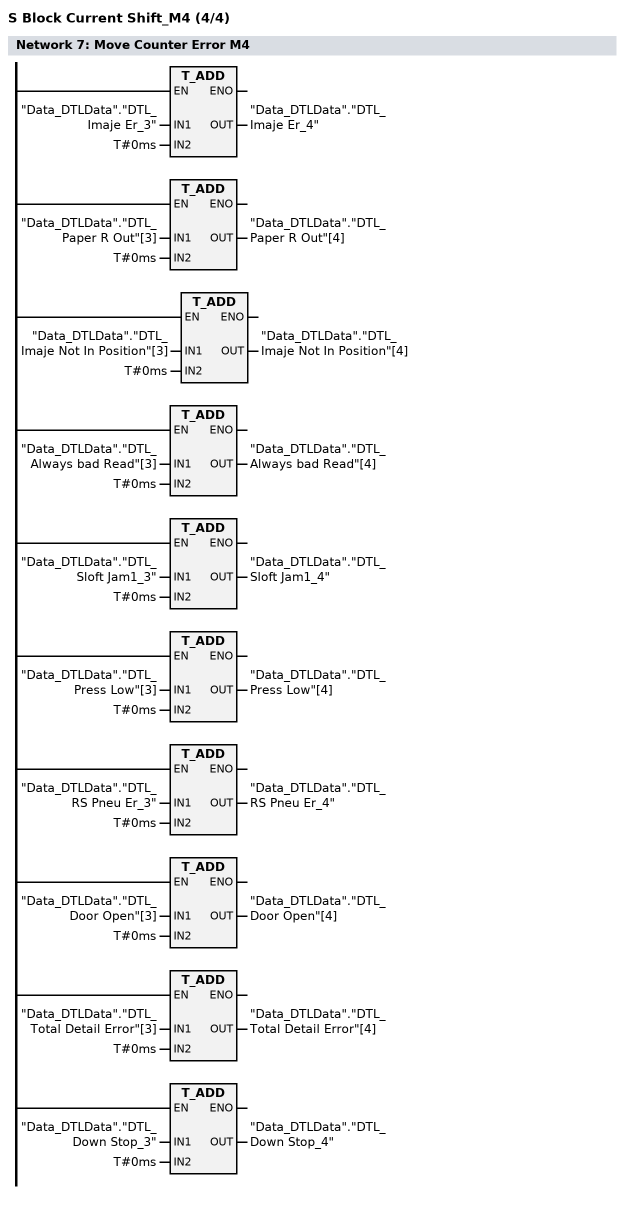
   "Data_DTLData"."DTL_Imaje Er_4" := T_ADD(IN1 := "Data_DTLData"."DTL_Imaje Er_3", IN2 := T#0ms);
   "Data_DTLData"."DTL_Paper R Out"[4] := T_ADD(IN1 := "Data_DTLData"."DTL_Paper R Out"[3], IN2 := T#0ms);
   "Data_DTLData"."DTL_Imaje Not In Position"[4] := T_ADD(IN1 := "Data_DTLData"."DTL_Imaje Not In Position"[3],
                           IN2 := T#0ms);
   "Data_DTLData"."DTL_Always bad Read"[4] := T_ADD(IN1 := "Data_DTLData"."DTL_Always bad Read"[3],
                           IN2 := T#0ms);
   "Data_DTLData"."DTL_Sloft Jam1_4" := T_ADD(IN1 := "Data_DTLData"."DTL_Sloft Jam1_3", IN2 := T#0ms);
   "Data_DTLData"."DTL_Press Low"[4] := T_ADD(IN1 := "Data_DTLData"."DTL_Press Low"[3], IN2 := T#0ms);
   "Data_DTLData"."DTL_RS Pneu Er_4" := T_ADD(IN1 := "Data_DTLData"."DTL_RS Pneu Er_3", IN2 := T#0ms);
   "Data_DTLData"."DTL_Door Open"[4] := T_ADD(IN1 := "Data_DTLData"."DTL_Door Open"[3], IN2 := T#0ms);
   "Data_DTLData"."DTL_Total Detail Error"[4] := T_ADD(IN1 := "Data_DTLData"."DTL_Total Detail Error"[3],
                           IN2 := T#0ms);
   "Data_DTLData"."DTL_Down Stop_4" := T_ADD(IN1 := "Data_DTLData"."DTL_Down Stop_3", IN2 := T#0ms);
END_REGION
END_FUNCTION_BLOCK

FUNCTION_BLOCK "S Block Current Shift_M5"   // FB14, LAD
{ S7_Optimized_Access := 'TRUE' }
VERSION : 0.1
BEGIN

REGION Network 1: Move Date Time M5
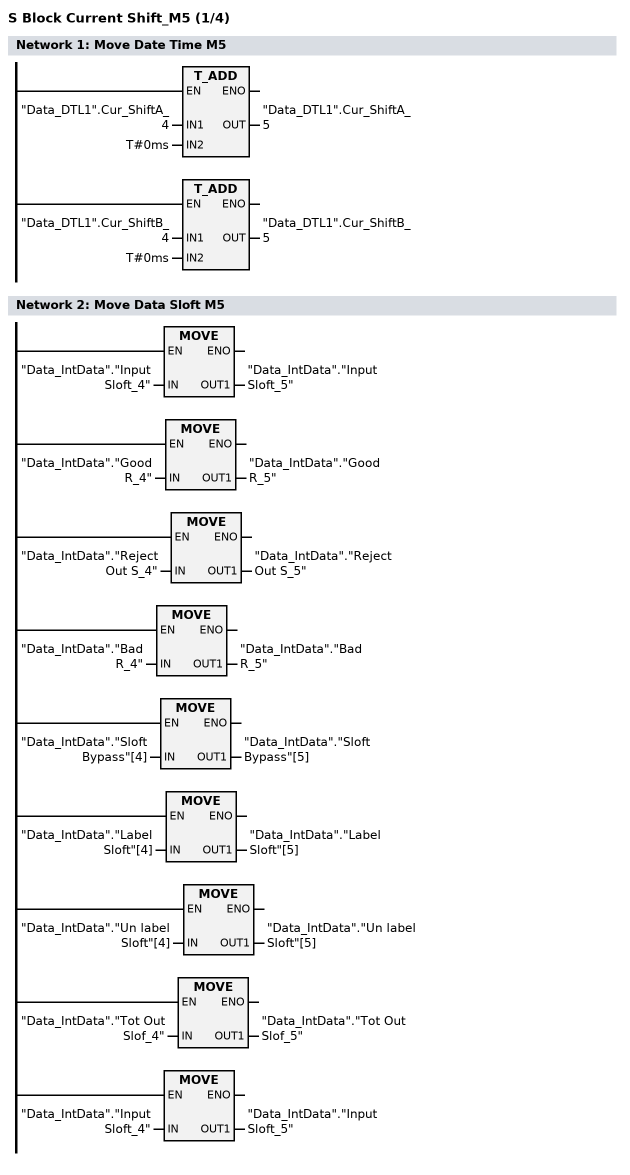
   "Data_DTL1".Cur_ShiftA_5 := T_ADD(IN1 := "Data_DTL1".Cur_ShiftA_4, IN2 := T#0ms);
   "Data_DTL1".Cur_ShiftB_5 := T_ADD(IN1 := "Data_DTL1".Cur_ShiftB_4, IN2 := T#0ms);
END_REGION

REGION Network 2: Move Data Sloft M5
   RUNG wire#powerrail
      { S7_GenerateENO := "TRUE" } Move(in := "Data_IntData"."Input Sloft_4", out1 => "Data_IntData"."Input Sloft_5")
   END_RUNG
   RUNG wire#powerrail
      { S7_GenerateENO := "TRUE" } Move(in := "Data_IntData"."Good R_4", out1 => "Data_IntData"."Good R_5")
   END_RUNG
   RUNG wire#powerrail
      { S7_GenerateENO := "TRUE" } Move(in := "Data_IntData"."Reject Out S_4", out1 => "Data_IntData"."Reject Out S_5")
   END_RUNG
   RUNG wire#powerrail
      { S7_GenerateENO := "TRUE" } Move(in := "Data_IntData"."Bad R_4", out1 => "Data_IntData"."Bad R_5")
   END_RUNG
   RUNG wire#powerrail
      { S7_GenerateENO := "TRUE" } Move(in := "Data_IntData"."Sloft Bypass"[4], out1 => "Data_IntData"."Sloft Bypass"[5])
   END_RUNG
   RUNG wire#powerrail
      { S7_GenerateENO := "TRUE" } Move(in := "Data_IntData"."Label Sloft"[4], out1 => "Data_IntData"."Label Sloft"[5])
   END_RUNG
   RUNG wire#powerrail
      { S7_GenerateENO := "TRUE" } Move(in := "Data_IntData"."Un label Sloft"[4], out1 => "Data_IntData"."Un label Sloft"[5])
   END_RUNG
   RUNG wire#powerrail
      { S7_GenerateENO := "TRUE" } Move(in := "Data_IntData"."Tot Out Slof_4", out1 => "Data_IntData"."Tot Out Slof_5")
   END_RUNG
   RUNG wire#powerrail
      { S7_GenerateENO := "TRUE" } Move(in := "Data_IntData"."Input Sloft_4", out1 => "Data_IntData"."Input Sloft_5")
   END_RUNG
   // the same network as SCL:
   "Data_IntData"."Input Sloft_5" := "Data_IntData"."Input Sloft_4";
   "Data_IntData"."Good R_5" := "Data_IntData"."Good R_4";
   "Data_IntData"."Reject Out S_5" := "Data_IntData"."Reject Out S_4";
   "Data_IntData"."Bad R_5" := "Data_IntData"."Bad R_4";
   "Data_IntData"."Sloft Bypass"[5] := "Data_IntData"."Sloft Bypass"[4];
   "Data_IntData"."Label Sloft"[5] := "Data_IntData"."Label Sloft"[4];
   "Data_IntData"."Un label Sloft"[5] := "Data_IntData"."Un label Sloft"[4];
   "Data_IntData"."Tot Out Slof_5" := "Data_IntData"."Tot Out Slof_4";
   "Data_IntData"."Input Sloft_5" := "Data_IntData"."Input Sloft_4";
END_REGION

REGION Network 3: Move Data Sloft Trigger & Aplicator M5
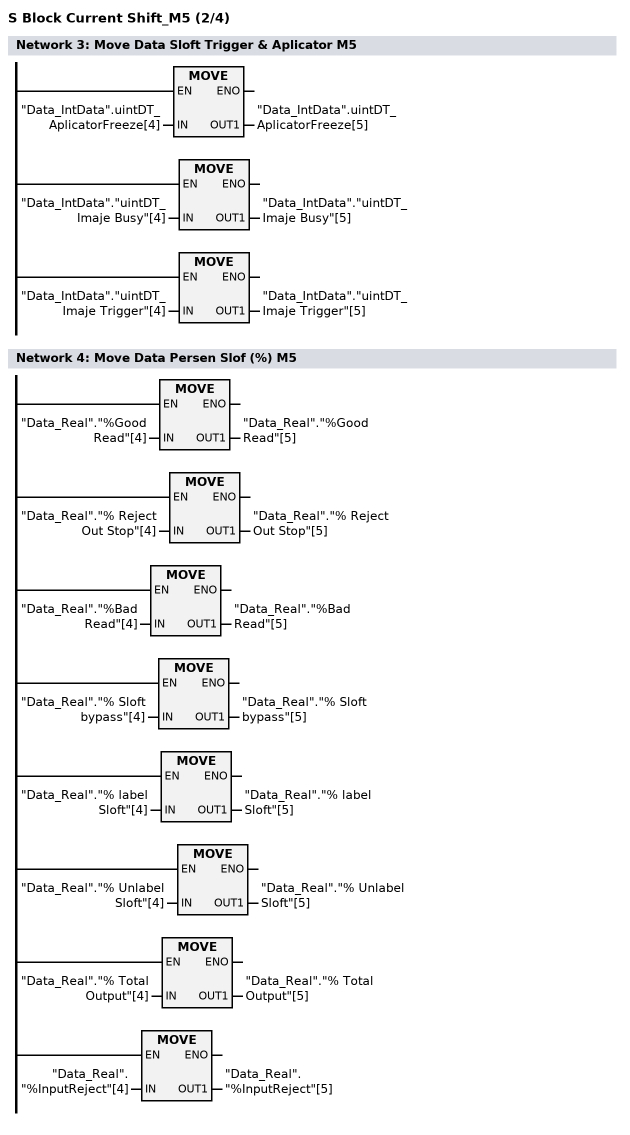
   RUNG wire#powerrail
      { S7_GenerateENO := "TRUE" } Move(in := "Data_IntData".uintDT_AplicatorFreeze[4], out1 => "Data_IntData".uintDT_AplicatorFreeze[5])
   END_RUNG
   RUNG wire#powerrail
      { S7_GenerateENO := "TRUE" } Move(in := "Data_IntData"."uintDT_Imaje Busy"[4], out1 => "Data_IntData"."uintDT_Imaje Busy"[5])
   END_RUNG
   RUNG wire#powerrail
      { S7_GenerateENO := "TRUE" } Move(in := "Data_IntData"."uintDT_Imaje Trigger"[4], out1 => "Data_IntData"."uintDT_Imaje Trigger"[5])
   END_RUNG
   // the same network as SCL:
   "Data_IntData".uintDT_AplicatorFreeze[5] := "Data_IntData".uintDT_AplicatorFreeze[4];
   "Data_IntData"."uintDT_Imaje Busy"[5] := "Data_IntData"."uintDT_Imaje Busy"[4];
   "Data_IntData"."uintDT_Imaje Trigger"[5] := "Data_IntData"."uintDT_Imaje Trigger"[4];
END_REGION

REGION Network 4: Move Data Persen Slof (%) M5
   RUNG wire#powerrail
      { S7_GenerateENO := "TRUE" } Move(in := "Data_Real"."%Good Read"[4], out1 => "Data_Real"."%Good Read"[5])
   END_RUNG
   RUNG wire#powerrail
      { S7_GenerateENO := "TRUE" } Move(in := "Data_Real"."% Reject Out Stop"[4], out1 => "Data_Real"."% Reject Out Stop"[5])
   END_RUNG
   RUNG wire#powerrail
      { S7_GenerateENO := "TRUE" } Move(in := "Data_Real"."%Bad Read"[4], out1 => "Data_Real"."%Bad Read"[5])
   END_RUNG
   RUNG wire#powerrail
      { S7_GenerateENO := "TRUE" } Move(in := "Data_Real"."% Sloft bypass"[4], out1 => "Data_Real"."% Sloft bypass"[5])
   END_RUNG
   RUNG wire#powerrail
      { S7_GenerateENO := "TRUE" } Move(in := "Data_Real"."% label Sloft"[4], out1 => "Data_Real"."% label Sloft"[5])
   END_RUNG
   RUNG wire#powerrail
      { S7_GenerateENO := "TRUE" } Move(in := "Data_Real"."% Unlabel Sloft"[4], out1 => "Data_Real"."% Unlabel Sloft"[5])
   END_RUNG
   RUNG wire#powerrail
      { S7_GenerateENO := "TRUE" } Move(in := "Data_Real"."% Total Output"[4], out1 => "Data_Real"."% Total Output"[5])
   END_RUNG
   RUNG wire#powerrail
      { S7_GenerateENO := "TRUE" } Move(in := "Data_Real"."%InputReject"[4], out1 => "Data_Real"."%InputReject"[5])
   END_RUNG
   // the same network as SCL:
   "Data_Real"."%Good Read"[5] := "Data_Real"."%Good Read"[4];
   "Data_Real"."% Reject Out Stop"[5] := "Data_Real"."% Reject Out Stop"[4];
   "Data_Real"."%Bad Read"[5] := "Data_Real"."%Bad Read"[4];
   "Data_Real"."% Sloft bypass"[5] := "Data_Real"."% Sloft bypass"[4];
   "Data_Real"."% label Sloft"[5] := "Data_Real"."% label Sloft"[4];
   "Data_Real"."% Unlabel Sloft"[5] := "Data_Real"."% Unlabel Sloft"[4];
   "Data_Real"."% Total Output"[5] := "Data_Real"."% Total Output"[4];
   "Data_Real"."%InputReject"[5] := "Data_Real"."%InputReject"[4];
END_REGION

REGION Network 5: Move Data Time Mesin M5
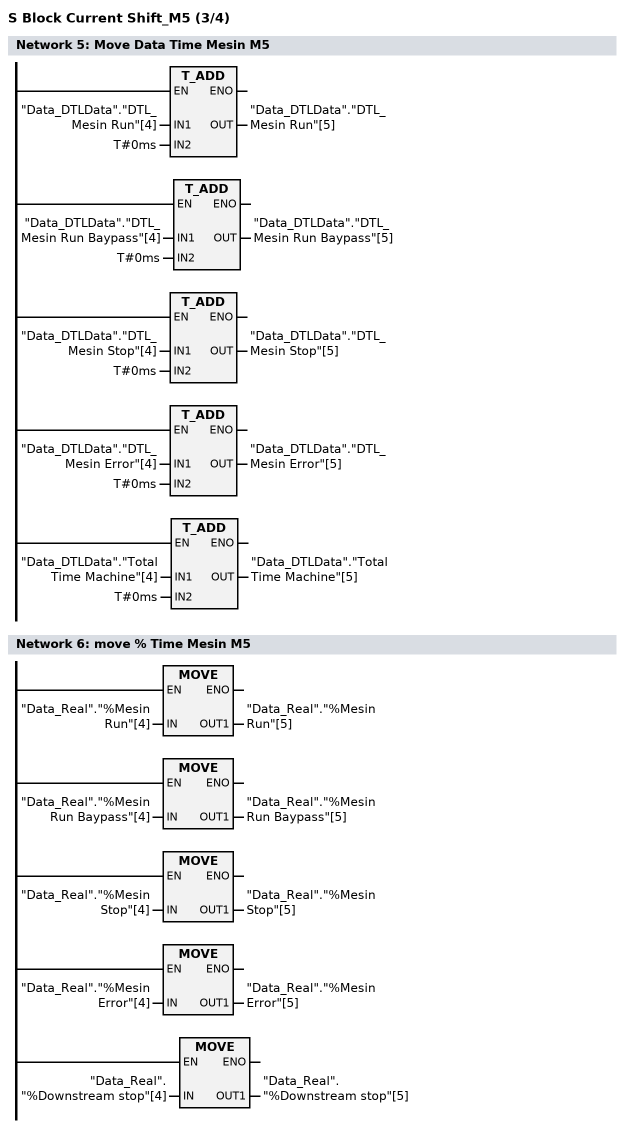
   "Data_DTLData"."DTL_Mesin Run"[5] := T_ADD(IN1 := "Data_DTLData"."DTL_Mesin Run"[4], IN2 := T#0ms);
   "Data_DTLData"."DTL_Mesin Run Baypass"[5] := T_ADD(IN1 := "Data_DTLData"."DTL_Mesin Run Baypass"[4],
                           IN2 := T#0ms);
   "Data_DTLData"."DTL_Mesin Stop"[5] := T_ADD(IN1 := "Data_DTLData"."DTL_Mesin Stop"[4], IN2 := T#0ms);
   "Data_DTLData"."DTL_Mesin Error"[5] := T_ADD(IN1 := "Data_DTLData"."DTL_Mesin Error"[4], IN2 := T#0ms);
   "Data_DTLData"."Total Time Machine"[5] := T_ADD(IN1 := "Data_DTLData"."Total Time Machine"[4], IN2 := T#0ms);
END_REGION

REGION Network 6: move % Time Mesin M5
   RUNG wire#powerrail
      { S7_GenerateENO := "TRUE" } Move(in := "Data_Real"."%Mesin Run"[4], out1 => "Data_Real"."%Mesin Run"[5])
   END_RUNG
   RUNG wire#powerrail
      { S7_GenerateENO := "TRUE" } Move(in := "Data_Real"."%Mesin Run Baypass"[4], out1 => "Data_Real"."%Mesin Run Baypass"[5])
   END_RUNG
   RUNG wire#powerrail
      { S7_GenerateENO := "TRUE" } Move(in := "Data_Real"."%Mesin Stop"[4], out1 => "Data_Real"."%Mesin Stop"[5])
   END_RUNG
   RUNG wire#powerrail
      { S7_GenerateENO := "TRUE" } Move(in := "Data_Real"."%Mesin Error"[4], out1 => "Data_Real"."%Mesin Error"[5])
   END_RUNG
   RUNG wire#powerrail
      { S7_GenerateENO := "TRUE" } Move(in := "Data_Real"."%Downstream stop"[4], out1 => "Data_Real"."%Downstream stop"[5])
   END_RUNG
   // the same network as SCL:
   "Data_Real"."%Mesin Run"[5] := "Data_Real"."%Mesin Run"[4];
   "Data_Real"."%Mesin Run Baypass"[5] := "Data_Real"."%Mesin Run Baypass"[4];
   "Data_Real"."%Mesin Stop"[5] := "Data_Real"."%Mesin Stop"[4];
   "Data_Real"."%Mesin Error"[5] := "Data_Real"."%Mesin Error"[4];
   "Data_Real"."%Downstream stop"[5] := "Data_Real"."%Downstream stop"[4];
END_REGION

REGION Network 7: Move Counter Error M5
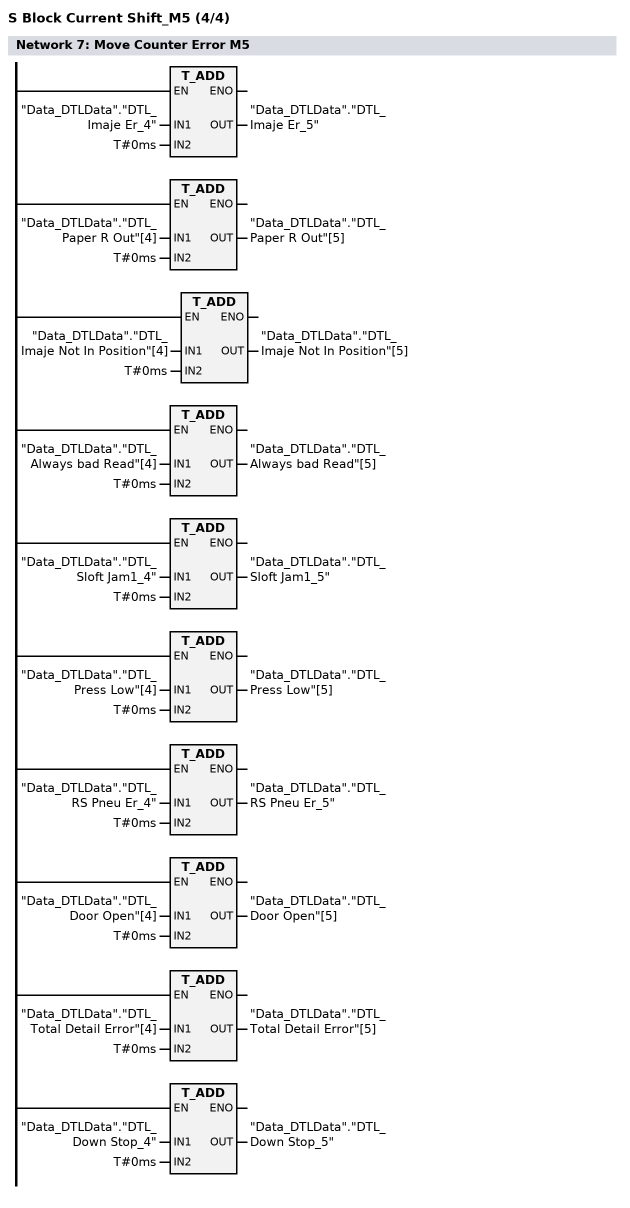
   "Data_DTLData"."DTL_Imaje Er_5" := T_ADD(IN1 := "Data_DTLData"."DTL_Imaje Er_4", IN2 := T#0ms);
   "Data_DTLData"."DTL_Paper R Out"[5] := T_ADD(IN1 := "Data_DTLData"."DTL_Paper R Out"[4], IN2 := T#0ms);
   "Data_DTLData"."DTL_Imaje Not In Position"[5] := T_ADD(IN1 := "Data_DTLData"."DTL_Imaje Not In Position"[4],
                           IN2 := T#0ms);
   "Data_DTLData"."DTL_Always bad Read"[5] := T_ADD(IN1 := "Data_DTLData"."DTL_Always bad Read"[4],
                           IN2 := T#0ms);
   "Data_DTLData"."DTL_Sloft Jam1_5" := T_ADD(IN1 := "Data_DTLData"."DTL_Sloft Jam1_4", IN2 := T#0ms);
   "Data_DTLData"."DTL_Press Low"[5] := T_ADD(IN1 := "Data_DTLData"."DTL_Press Low"[4], IN2 := T#0ms);
   "Data_DTLData"."DTL_RS Pneu Er_5" := T_ADD(IN1 := "Data_DTLData"."DTL_RS Pneu Er_4", IN2 := T#0ms);
   "Data_DTLData"."DTL_Door Open"[5] := T_ADD(IN1 := "Data_DTLData"."DTL_Door Open"[4], IN2 := T#0ms);
   "Data_DTLData"."DTL_Total Detail Error"[5] := T_ADD(IN1 := "Data_DTLData"."DTL_Total Detail Error"[4],
                           IN2 := T#0ms);
   "Data_DTLData"."DTL_Down Stop_5" := T_ADD(IN1 := "Data_DTLData"."DTL_Down Stop_4", IN2 := T#0ms);
END_REGION
END_FUNCTION_BLOCK

FUNCTION_BLOCK "AddReject2"   // FB15, SCL
{ S7_Optimized_Access := 'TRUE' }
VERSION : 0.1
   VAR_INPUT
      Sensor1 : Bool;
      Sensor2 : Bool;
      Sensor3 : Bool;
      Reedswicth1 : Bool;
      Reedswicth2 : Bool;
      BypassRS_AddRej : Bool;
      BypassRS_All_RS : Bool;
      PT_Timer_S1On : Time;
      PT_Timer_S1Off : Time;
      PT_Timer_S2On : Time;
      PT_Timer_S2Off : Time;
      PT_Timer_S3On : Time;
      PT_Timer_S3Off : Time;
      PT_Timer_DelayReject : Time;
      PT_Timer_DelayNonReject : Time;
   END_VAR
   VAR_OUTPUT
      Pneumatic1 : Bool;
      Pneumatic2 : Bool;
      Countaddrej : Time;
   END_VAR
   VAR
      SeqIndexReject : UInt;
      SeqIndexNonReject : UInt;
      FlagReject : Bool;
      FlagNonReject : Bool;
      FlagPneumatic : Bool;
      FlagSensor1 : Bool;
      FlagSensor2 : Bool;
      FlagSensor3 : Bool;
      FlagRS1Advance : Bool;
      FlagRS2Retract : Bool;
      RS1AdvanceError : Bool;
      RS2RetractError : Bool;
      AllRSAddRejectError : Bool;
      CountStop : Bool;
      InTimerDelayReject : Bool;
      InTimerDelaynonReject : Bool;
      InTimerErrorReject : Bool;
      InTimerErrorNonReject : Bool;
      InTimerRS1Error : Bool;
      InTimerRS2Error : Bool;
      R_TRIG_AddRejPSN1 : R_TRIG;
      F_TRIG_AddRejPSN1 : F_TRIG;
   END_VAR
BEGIN
   //Sensor 1
   "ttM_TimerAddRej1".TON(IN := #Sensor1,
                          PT := #PT_Timer_S1On);
   "tTM_TimerAddRej2".TON(IN := NOT #Sensor1,
                          PT := #PT_Timer_S1Off);
   IF "ttM_TimerAddRej1".Q THEN
       #FlagSensor1 := TRUE;
   END_IF;
   IF "tTM_TimerAddRej2".Q THEN
       #FlagSensor1 := FALSE;
   END_IF;

   //Sensor 2
   "tTM_TimerAddRej3".TON(IN := #Sensor2,
                          PT := #PT_Timer_S2On);
   "tTM_TimerAddRej4".TON(IN := NOT #Sensor2,
                          PT := #PT_Timer_S2Off);
   IF "tTM_TimerAddRej3".Q THEN
       #FlagSensor2 := TRUE;
   END_IF;
   IF "tTM_TimerAddRej4".Q THEN
       #FlagSensor2 := FALSE;
   END_IF;

   //Sensor 3
   "tTM_TimerAddRej5".TON(IN := #Sensor3,
                          PT := #PT_Timer_S3On);
   "tTM_TimerAddRej6".TON(IN := NOT #Sensor3,
                          PT := #PT_Timer_S3Off);
   IF "tTM_TimerAddRej5".Q THEN
       #FlagSensor3 := TRUE;
   END_IF;
   IF "tTM_TimerAddRej6".Q THEN
       #FlagSensor3 := FALSE;
   END_IF;

   //Reedswicth
   "tTM_TimerRS1_Adv".TON(IN := #InTimerRS1Error,
                          PT := T#1700ms);
   "tTM_TimerRS2_Ret".TON(IN := #InTimerRS2Error,
                          PT := T#1700ms);
   IF NOT #BypassRS_AddRej AND NOT #BypassRS_All_RS THEN
       //ReedSwicth Advance
       IF NOT #Pneumatic1 THEN
           #InTimerRS1Error := TRUE;
           "R_TRIG_RS1_Adv"(CLK := #Reedswicth1);
           IF #Reedswicth1 OR "R_TRIG_RS1_Adv".Q THEN
               #FlagRS1Advance := TRUE;
               #FlagRS2Retract := FALSE;
               #RS1AdvanceError := FALSE;
               #RS2RetractError := FALSE;
           ELSIF "tTM_TimerRS1_Adv".Q AND NOT #FlagRS1Advance THEN
               #FlagRS1Advance := FALSE;
               #FlagRS2Retract := FALSE;
               #RS1AdvanceError := TRUE;
               #RS2RetractError := FALSE;
           END_IF;
       ELSE
           #InTimerRS1Error := FALSE;
       END_IF;
       //ReeedSwicth Retract
       IF #Pneumatic2 THEN
           #InTimerRS2Error := TRUE;
           "R_TRIG_RS2_Ret"(CLK := #Reedswicth2);
           IF #Reedswicth2 OR "R_TRIG_RS2_Ret".Q THEN
               #FlagRS1Advance := FALSE;
               #FlagRS2Retract := TRUE;
               #RS1AdvanceError := FALSE;
               #RS2RetractError := FALSE;
           ELSIF "tTM_TimerRS2_Ret".Q AND NOT #FlagRS2Retract THEN
               #FlagRS1Advance := FALSE;
               #FlagRS2Retract := FALSE;
               #RS1AdvanceError := FALSE;
               #RS2RetractError := TRUE;
           END_IF;
       ELSE
           #InTimerRS2Error := FALSE;
       END_IF;
       //Error All ReedSwicth
       IF NOT #FlagRS1Advance AND NOT #FlagRS2Retract THEN
           "tTM_ErrorAllRSAddReject".TON(IN:=NOT #FlagRS1Advance AND NOT #FlagRS2Retract,
                                         PT:=T#3500ms);
           IF "tTM_ErrorAllRSAddReject".Q THEN
               IF #FlagSensor1 THEN
                   #Pneumatic1 := TRUE;
                   #Pneumatic2 := TRUE;
               ELSE
                   #Pneumatic1 := FALSE;
                   #Pneumatic2 := FALSE;
               END_IF;
               #AllRSAddRejectError := TRUE;
               #SeqIndexReject := 0;
               #SeqIndexNonReject := 0;
           END_IF;
       ELSE
           #AllRSAddRejectError := FALSE;
           "F_TRIG_AllRSAddrejError"(CLK:=#AllRSAddRejectError);
           IF "F_TRIG_AllRSAddrejError".Q THEN
               #SeqIndexReject := 1;
               #SeqIndexNonReject := 1;
           END_IF;
       END_IF;
   END_IF;

   //Reject Active
   IF #FlagSensor1 THEN
       IF NOT #AllRSAddRejectError THEN
           #SeqIndexNonReject := 1;
       END_IF;
       "tTM_DelayReject".TON(IN := #InTimerDelayReject,
                             PT := #PT_Timer_DelayReject);
       "tTM_ErrorReject".TON(IN := #InTimerErrorReject,
                             PT := T#2000ms);
       CASE #SeqIndexReject OF
           1:
               #InTimerErrorReject := FALSE;
               IF NOT #FlagSensor2 THEN
                   #Pneumatic1 := FALSE;
                   #Pneumatic2 := FALSE;
                   #SeqIndexReject := 10;
               ELSIF #FlagSensor2 THEN
                   IF "tTM_DelayReject".Q THEN
                       #Pneumatic1 := FALSE;
                       #Pneumatic2 := FALSE;
                       #SeqIndexReject := 10;
                   ELSE
                       #InTimerDelayReject := TRUE;
                   END_IF;
               END_IF;
           10:
               #InTimerDelayReject := FALSE;
               IF NOT #BypassRS_AddRej AND NOT #BypassRS_All_RS THEN
                   #SeqIndexReject := 20;
               ELSE
                   #SeqIndexReject := 1;
               END_IF;
           20:
               IF #FlagRS1Advance THEN
                   #SeqIndexReject := 1;
               ELSIF #RS1AdvanceError THEN
                   #Pneumatic1 := TRUE;
                   #Pneumatic2 := TRUE;
                   IF "tTM_ErrorReject".Q THEN
                       #SeqIndexReject := 1;
                   ELSE
                       #InTimerErrorReject := TRUE;
                   END_IF;
               END_IF;
           ELSE
               IF NOT #BypassRS_AddRej AND NOT #BypassRS_All_RS AND NOT #AllRSAddRejectError  THEN
                   #SeqIndexReject := 1;
               ELSE
                   #SeqIndexReject := 1;
               END_IF;
       END_CASE;
   END_IF;

   //Reject Start Non Active 
   IF NOT #FlagSensor1  THEN
       IF NOT #AllRSAddRejectError THEN
           #SeqIndexReject := 1;
       END_IF;
       "tTM_DelayNonReject".TON(IN := #InTimerDelaynonReject,
                                PT := #PT_Timer_DelayNonReject);
       "tTM_ErrorNonReject".TON(IN := #InTimerErrorNonReject,
                                PT := T#2000ms);
       CASE #SeqIndexNonReject OF
           1:
               #InTimerErrorNonReject := FALSE;
               IF NOT #FlagSensor3 THEN
                   #Pneumatic1 := TRUE;
                   #Pneumatic2 := TRUE;
                   #SeqIndexNonReject := 10;
               ELSIF #FlagSensor3 THEN
                   IF "tTM_DelayNonReject".Q THEN
                       #Pneumatic1 := TRUE;
                       #Pneumatic2 := TRUE;
                       #SeqIndexNonReject := 10;
                   ELSE
                       #InTimerDelaynonReject := TRUE;
                   END_IF;
               END_IF;
           10:
               #InTimerDelaynonReject := FALSE;
               IF NOT #BypassRS_AddRej AND NOT #BypassRS_All_RS THEN
                   #SeqIndexNonReject := 20;
               ELSE
                   #SeqIndexNonReject := 1;
               END_IF;
           20:
               IF #FlagRS2Retract THEN
                   #SeqIndexNonReject := 1;
               ELSIF #RS2RetractError THEN
                   #Pneumatic1 := FALSE;
                   #Pneumatic2 := FALSE;
                   IF "tTM_ErrorNonReject".Q THEN
                       #SeqIndexNonReject := 1;
                   ELSE
                       #InTimerErrorNonReject := TRUE;
                   END_IF;
               END_IF;
           ELSE
               IF NOT #BypassRS_AddRej AND NOT #BypassRS_All_RS AND NOT #AllRSAddRejectError THEN
                   #SeqIndexNonReject := 1;
               ELSE
                   #SeqIndexNonReject := 1;
               END_IF;
       END_CASE;
   END_IF;

   #R_TRIG_AddRejPSN1(CLK:=#FlagSensor1);
   #F_TRIG_AddRejPSN1(CLK:=#FlagSensor1);
   IF NOT #AllRSAddRejectError THEN
       IF #R_TRIG_AddRejPSN1.Q THEN
           #SeqIndexReject := 1;
       END_IF;
       IF #F_TRIG_AddRejPSN1.Q THEN
           #SeqIndexNonReject := 1;
       END_IF;
   END_IF;

   "tTM_CountAddReject".TON(IN:=#Sensor1,
                            PT:=T#5000ms);
   IF "tTM_CountAddReject".ET <>T#0ms THEN
       #Countaddrej :="tTM_CountAddReject".ET;
   ELSIF #CountStop THEN
       #Countaddrej := T#0ms;
   END_IF;


   //Error All ReedSwicth

   //Reject Active
   (*IF #FlagSensor1 THEN
     IF NOT #FlagSensor2 THEN
       #Pneumatic1 := FALSE;
       #Pneumatic2 := FALSE;
       #FlagPneumatic := FALSE;
     END_IF;
   END_IF;
   //Reject Start Non Active 
   IF NOT #FlagSensor1 THEN
       IF NOT #FlagSensor3 THEN
           #Pneumatic1 := TRUE;
           #Pneumatic2 := TRUE;
           #FlagPneumatic := TRUE;
       END_IF;
   END_IF;

   CASE #SeqIndex OF
       0:
           #RS1Error := FALSE;
           #RS2Error := FALSE;
           //Reject Start Active
           IF #FlagSensor1 AND NOT #RejectActive THEN
               #SeqIndex := 5;
           END_IF;
           //Reject Start Non Active 
           IF NOT #FlagSensor1 AND #RejectActive THEN
               #SeqIndex := 10;
           END_IF;
       5: //Reject Active
           IF NOT #FlagSensor2 THEN
               #Pneumatic1 := FALSE;
               #Pneumatic2 := FALSE;
               #FlagPneumatic := FALSE;
               #SeqIndex := 15;
           END_IF;
       10: //Reject Non Active
           IF NOT #FlagSensor3 THEN
               #Pneumatic1 := TRUE;
               #Pneumatic2 := TRUE;
               #FlagPneumatic := TRUE;
               #SeqIndex := 20;
           END_IF;
       15: // Active Finish
           IF #BypassRS_AddRej OR #BypassRS_All_RS THEN
               #RejectActive := TRUE;
               #SeqIndex := 0;
           ELSIF NOT #BypassRS_AddRej AND NOT #BypassRS_All_RS THEN
               IF #FlagRS1 THEN
                   #RejectActive := TRUE;
                   #SeqIndex := 0;
               ELSIF #RS1Error THEN
                   #Pneumatic1 := TRUE;
                   #Pneumatic2 := TRUE;
                   #FlagPneumatic := TRUE;
                   #RejectActive := FALSE;
                   #SeqIndex := 0;
               END_IF;
           END_IF;
       20: //Cek Non Active Finish
           IF #BypassRS_AddRej OR #BypassRS_All_RS THEN
               #RejectActive := FALSE;
               #SeqIndex := 0;
           ELSIF NOT #BypassRS_AddRej AND NOT #BypassRS_All_RS THEN
               IF #FlagRS2 THEN
                   #RejectActive := FALSE;
                   #SeqIndex := 0;
               ELSIF #RS2Error THEN
                   #Pneumatic1 := FALSE;
                   #Pneumatic2 := FALSE;
                   #FlagPneumatic := FALSE;
                   #RejectActive := TRUE;
                   #SeqIndex := 0;
               END_IF;
           END_IF;
       END_CASE;*)
END_FUNCTION_BLOCK

FUNCTION "RS 1 Pneumatic Pusher Advance" : Void   // FC1, LAD
{ S7_Optimized_Access := 'TRUE' }
VERSION : 0.1
BEGIN

REGION Network 1: Reed Switch Pneumatic 1 Advance Ready
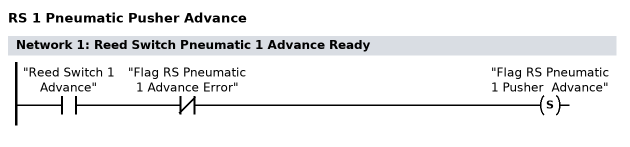
   RUNG wire#powerrail
      Contact( "Reed Switch 1 Advance" )
      I_Contact( "Flag RS Pneumatic 1 Advance Error" )
      S_Coil( "Flag RS Pneumatic 1 Pusher  Advance" )
   END_RUNG
   // the same network as SCL:
   IF "Reed Switch 1 Advance" AND NOT "Flag RS Pneumatic 1 Advance Error" THEN
       "Flag RS Pneumatic 1 Pusher  Advance" := TRUE;
   END_IF;
END_REGION
END_FUNCTION

FUNCTION "RS 2 Pneumatic Pusher Retract" : Void   // FC2, LAD
{ S7_Optimized_Access := 'TRUE' }
VERSION : 0.1
BEGIN

REGION Network 1: Reed Switch Pneumatic 1 Upper Ready
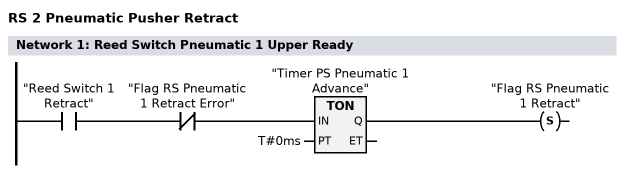
   "Timer PS Pneumatic 1 Advance".TON(IN := "Reed Switch 1 Retract" AND NOT "Flag RS Pneumatic 1 Retract Error",
                           PT := T#0ms);
   IF "Timer PS Pneumatic 1 Advance".Q THEN "Flag RS Pneumatic 1 Retract" := TRUE; END_IF;
END_REGION
END_FUNCTION

FUNCTION "RS 3 Pneumatic 3 Up" : Void   // FC3, LAD
{ S7_Optimized_Access := 'TRUE' }
VERSION : 0.1
BEGIN

REGION Network 1: Reed Switch Pneumatic 3 Up Ready
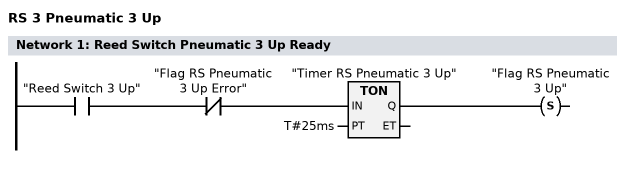
   "Timer RS Pneumatic 3 Up".TON(IN := "Reed Switch 3 Up" AND NOT "Flag RS Pneumatic 3 Up Error", PT := T#25ms);
   IF "Timer RS Pneumatic 3 Up".Q THEN "Flag RS Pneumatic 3 Up" := TRUE; END_IF;
END_REGION
END_FUNCTION

FUNCTION "RS 4 Pneumatic 3 Down" : Void   // FC4, LAD
{ S7_Optimized_Access := 'TRUE' }
VERSION : 0.1
BEGIN

REGION Network 1: Reed Switch Pneumatic 3 Down Ready
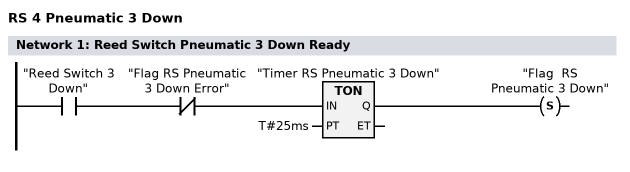
   "Timer RS Pneumatic 3 Down".TON(IN := "Reed Switch 3 Down" AND NOT "Flag RS Pneumatic 3 Down Error",
                           PT := T#25ms);
   IF "Timer RS Pneumatic 3 Down".Q THEN "Flag  RS Pneumatic 3 Down" := TRUE; END_IF;
END_REGION
END_FUNCTION

FUNCTION "RS 5 Pneumatic 4 Down" : Void   // FC5, LAD
{ S7_Optimized_Access := 'TRUE' }
VERSION : 0.1
BEGIN

REGION Network 1: Reed Switch Pneumatic 4 Down Ready
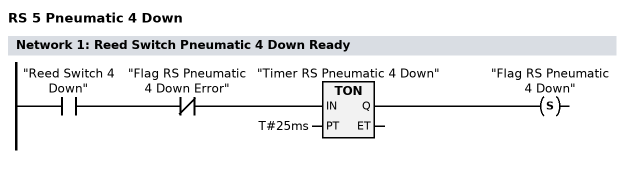
   "Timer RS Pneumatic 4 Down".TON(IN := "Reed Switch 4 Down" AND NOT "Flag RS Pneumatic 4 Down Error",
                           PT := T#25ms);
   IF "Timer RS Pneumatic 4 Down".Q THEN "Flag RS Pneumatic 4 Down" := TRUE; END_IF;
END_REGION
END_FUNCTION

FUNCTION "RS 6 Pneumatic 4 Up" : Void   // FC6, LAD
{ S7_Optimized_Access := 'TRUE' }
VERSION : 0.1
BEGIN

REGION Network 1: Reed Switch Pneumatic 4 Up Ready
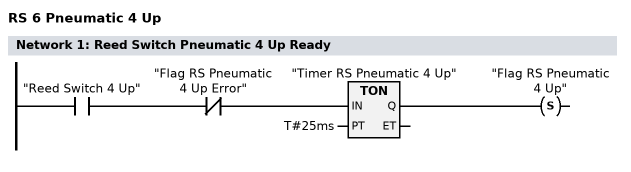
   "Timer RS Pneumatic 4 Up".TON(IN := "Reed Switch 4 Up" AND NOT "Flag RS Pneumatic 4 Up Error", PT := T#25ms);
   IF "Timer RS Pneumatic 4 Up".Q THEN "Flag RS Pneumatic 4 Up" := TRUE; END_IF;
END_REGION
END_FUNCTION

FUNCTION "RS 7 Pneumatic 5 Advance" : Void   // FC7, LAD
{ S7_Optimized_Access := 'TRUE' }
VERSION : 0.1
BEGIN

REGION Network 1: Reed Switch Pneumatic 5 Advance Ready
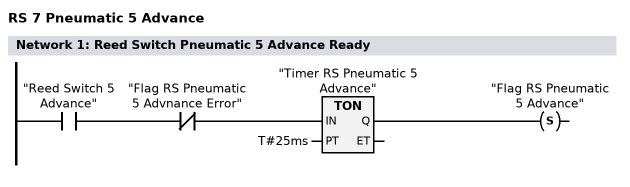
   "Timer RS Pneumatic 5 Advance".TON(IN := "Reed Switch 5 Advance" AND NOT "Flag RS Pneumatic 5 Advnance Error",
                           PT := T#25ms);
   IF "Timer RS Pneumatic 5 Advance".Q THEN "Flag RS Pneumatic 5 Advance" := TRUE; END_IF;
END_REGION
END_FUNCTION

FUNCTION "RS 8 Pneumatic 5 Retract" : Void   // FC8, LAD
{ S7_Optimized_Access := 'TRUE' }
VERSION : 0.1
BEGIN

REGION Network 1: Reed Switch Pneumatic 5 Retract Ready
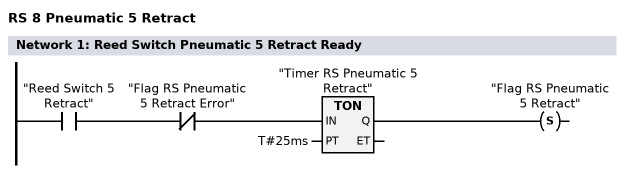
   "Timer RS Pneumatic 5 Retract".TON(IN := "Reed Switch 5 Retract" AND NOT "Flag RS Pneumatic 5 Retract Error",
                           PT := T#25ms);
   IF "Timer RS Pneumatic 5 Retract".Q THEN "Flag RS Pneumatic 5 Retract" := TRUE; END_IF;
END_REGION
END_FUNCTION

ORGANIZATION_BLOCK "Main"   // OB1, LAD, ProgramCycle
TITLE = "Main Program Sweep (Cycle)"
{ S7_Optimized_Access := 'TRUE' }
VERSION : 0.1
   VAR_TEMP   // added for the SCL form of the ladder/FBD networks
      _w1 : Bool;
      _w2 : Bool;
      _w3 : Bool;
      _w4 : Bool;
      _w5 : Bool;
   END_VAR
BEGIN

REGION Network 1: Machine Stand by
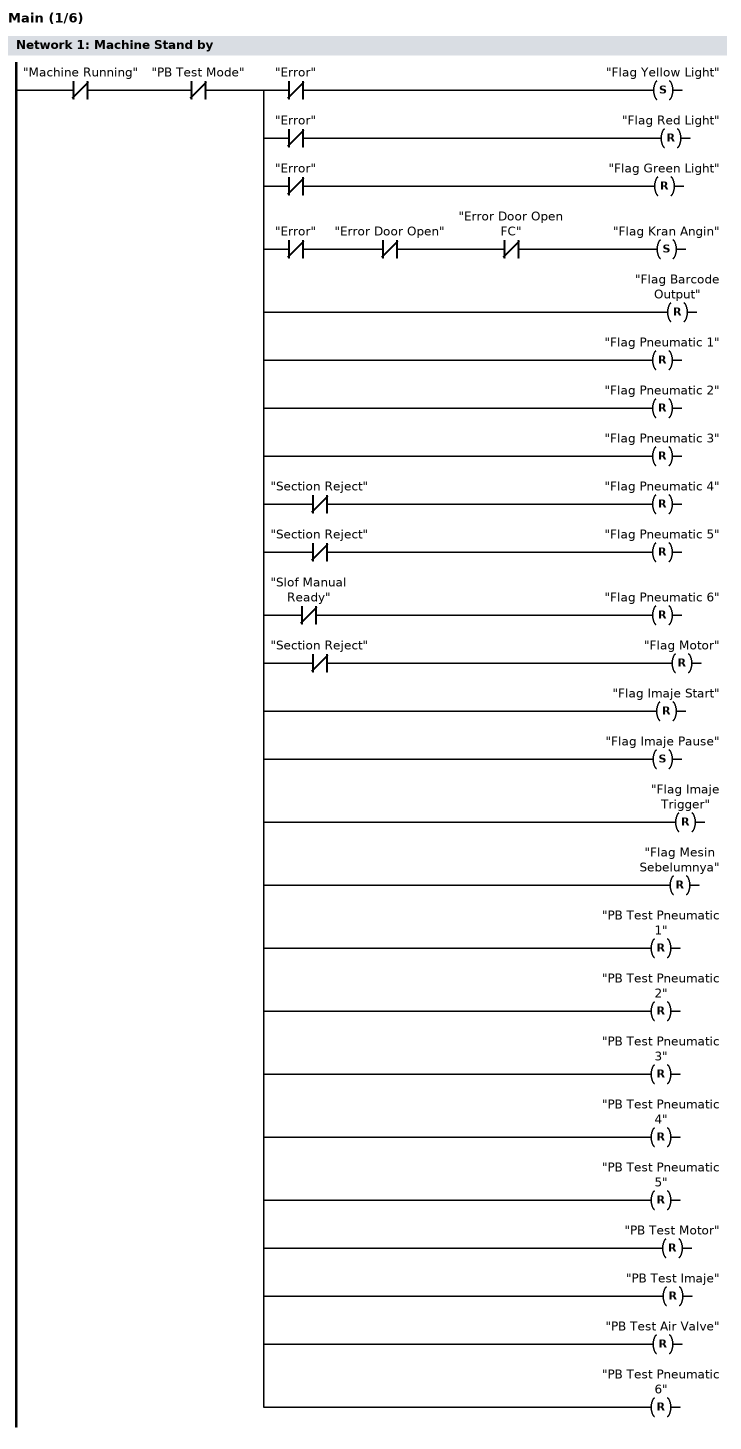
   RUNG wire#powerrail
      I_Contact( "Machine Running" )
      I_Contact( "PB Test Mode" )
      wire#w1
      I_Contact( "Error" )
      S_Coil( "Flag Yellow Light" )
   END_RUNG
   RUNG wire#w1
      I_Contact( "Error" )
      R_Coil( "Flag Red Light" )
   END_RUNG
   RUNG wire#w1
      I_Contact( "Error" )
      R_Coil( "Flag Green Light" )
   END_RUNG
   RUNG wire#w1
      I_Contact( "Error" )
      I_Contact( "Error Door Open" )
      I_Contact( "Error Door Open FC" )
      S_Coil( "Flag Kran Angin" )
   END_RUNG
   RUNG wire#w1
      R_Coil( "Flag Barcode Output" )
   END_RUNG
   RUNG wire#w1
      R_Coil( "Flag Pneumatic 1" )
   END_RUNG
   RUNG wire#w1
      R_Coil( "Flag Pneumatic 2" )
   END_RUNG
   RUNG wire#w1
      R_Coil( "Flag Pneumatic 3" )
   END_RUNG
   RUNG wire#w1
      I_Contact( "Section Reject" )
      R_Coil( "Flag Pneumatic 4" )
   END_RUNG
   RUNG wire#w1
      I_Contact( "Section Reject" )
      R_Coil( "Flag Pneumatic 5" )
   END_RUNG
   RUNG wire#w1
      I_Contact( "Slof Manual Ready" )
      R_Coil( "Flag Pneumatic 6" )
   END_RUNG
   RUNG wire#w1
      I_Contact( "Section Reject" )
      R_Coil( "Flag Motor" )
   END_RUNG
   RUNG wire#w1
      R_Coil( "Flag Imaje Start" )
   END_RUNG
   RUNG wire#w1
      S_Coil( "Flag Imaje Pause" )
   END_RUNG
   RUNG wire#w1
      R_Coil( "Flag Imaje Trigger" )
   END_RUNG
   RUNG wire#w1
      R_Coil( "Flag Mesin Sebelumnya" )
   END_RUNG
   RUNG wire#w1
      R_Coil( "PB Test Pneumatic 1" )
   END_RUNG
   RUNG wire#w1
      R_Coil( "PB Test Pneumatic 2" )
   END_RUNG
   RUNG wire#w1
      R_Coil( "PB Test Pneumatic 3" )
   END_RUNG
   RUNG wire#w1
      R_Coil( "PB Test Pneumatic 4" )
   END_RUNG
   RUNG wire#w1
      R_Coil( "PB Test Pneumatic 5" )
   END_RUNG
   RUNG wire#w1
      R_Coil( "PB Test Motor" )
   END_RUNG
   RUNG wire#w1
      R_Coil( "PB Test Imaje" )